REGION Network 14
   RUNG wire#powerrail
      #"2#柴油泵电动阀"(READY := "2#柴油泵电动蝶阀备妥", RUN := "2#柴油泵电动蝶阀运行", FAULT := "2#柴油泵电动蝶阀故障", OPEN_END := "2#柴油泵电动蝶阀开到位", CLOSE_END := "2#柴油泵电动蝶阀关到位", HMI_OPEN :=, HMI_CLOSE :=, MA :=, AUTO_OPEN :=, AUTO_CLOSE :=, QD_OPEN := "2#柴油泵电动阀开", QD_CLOSE := "2#柴油泵电动阀关")
   END_RUNG
   // the same network as SCL:
   #"2#柴油泵电动阀"(READY := "2#柴油泵电动蝶阀备妥",   // "阀门_MODEL"
               RUN := "2#柴油泵电动蝶阀运行",
               FAULT := "2#柴油泵电动蝶阀故障",
               OPEN_END := "2#柴油泵电动蝶阀开到位",
               CLOSE_END := "2#柴油泵电动蝶阀关到位",
               QD_OPEN := "2#柴油泵电动阀开",
               QD_CLOSE := "2#柴油泵电动阀关");
END_REGION

REGION Network 15
   RUNG wire#powerrail
      #"1#浊环热水泵电动阀"(READY := "1#浊环热水电动蝶阀备妥", RUN := "1#浊环热水电动蝶阀运行", FAULT := "1#浊环热水电动蝶阀故障", OPEN_END := "1#浊环热水电动蝶阀开到位", CLOSE_END := "1#浊环热水电动蝶阀关到位", HMI_OPEN :=, HMI_CLOSE :=, MA :=, AUTO_OPEN :=, AUTO_CLOSE :=, QD_OPEN := "1#浊环热水泵电动阀开", QD_CLOSE := "1#浊环热水泵电动阀关")
   END_RUNG
   // the same network as SCL:
   #"1#浊环热水泵电动阀"(READY := "1#浊环热水电动蝶阀备妥",   // "阀门_MODEL"
                 RUN := "1#浊环热水电动蝶阀运行",
                 FAULT := "1#浊环热水电动蝶阀故障",
                 OPEN_END := "1#浊环热水电动蝶阀开到位",
                 CLOSE_END := "1#浊环热水电动蝶阀关到位",
                 QD_OPEN := "1#浊环热水泵电动阀开",
                 QD_CLOSE := "1#浊环热水泵电动阀关");
END_REGION

REGION Network 16
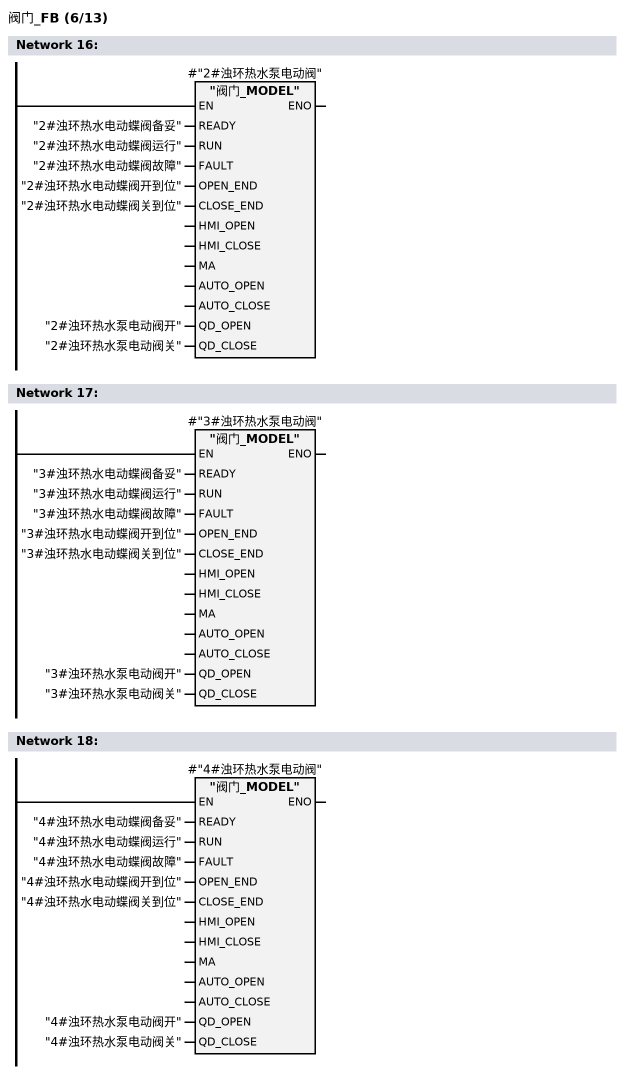
   RUNG wire#powerrail
      #"2#浊环热水泵电动阀"(READY := "2#浊环热水电动蝶阀备妥", RUN := "2#浊环热水电动蝶阀运行", FAULT := "2#浊环热水电动蝶阀故障", OPEN_END := "2#浊环热水电动蝶阀开到位", CLOSE_END := "2#浊环热水电动蝶阀关到位", HMI_OPEN :=, HMI_CLOSE :=, MA :=, AUTO_OPEN :=, AUTO_CLOSE :=, QD_OPEN := "2#浊环热水泵电动阀开", QD_CLOSE := "2#浊环热水泵电动阀关")
   END_RUNG
   // the same network as SCL:
   #"2#浊环热水泵电动阀"(READY := "2#浊环热水电动蝶阀备妥",   // "阀门_MODEL"
                 RUN := "2#浊环热水电动蝶阀运行",
                 FAULT := "2#浊环热水电动蝶阀故障",
                 OPEN_END := "2#浊环热水电动蝶阀开到位",
                 CLOSE_END := "2#浊环热水电动蝶阀关到位",
                 QD_OPEN := "2#浊环热水泵电动阀开",
                 QD_CLOSE := "2#浊环热水泵电动阀关");
END_REGION

REGION Network 17
   RUNG wire#powerrail
      #"3#浊环热水泵电动阀"(READY := "3#浊环热水电动蝶阀备妥", RUN := "3#浊环热水电动蝶阀运行", FAULT := "3#浊环热水电动蝶阀故障", OPEN_END := "3#浊环热水电动蝶阀开到位", CLOSE_END := "3#浊环热水电动蝶阀关到位", HMI_OPEN :=, HMI_CLOSE :=, MA :=, AUTO_OPEN :=, AUTO_CLOSE :=, QD_OPEN := "3#浊环热水泵电动阀开", QD_CLOSE := "3#浊环热水泵电动阀关")
   END_RUNG
   // the same network as SCL:
   #"3#浊环热水泵电动阀"(READY := "3#浊环热水电动蝶阀备妥",   // "阀门_MODEL"
                 RUN := "3#浊环热水电动蝶阀运行",
                 FAULT := "3#浊环热水电动蝶阀故障",
                 OPEN_END := "3#浊环热水电动蝶阀开到位",
                 CLOSE_END := "3#浊环热水电动蝶阀关到位",
                 QD_OPEN := "3#浊环热水泵电动阀开",
                 QD_CLOSE := "3#浊环热水泵电动阀关");
END_REGION

REGION Network 18
   RUNG wire#powerrail
      #"4#浊环热水泵电动阀"(READY := "4#浊环热水电动蝶阀备妥", RUN := "4#浊环热水电动蝶阀运行", FAULT := "4#浊环热水电动蝶阀故障", OPEN_END := "4#浊环热水电动蝶阀开到位", CLOSE_END := "4#浊环热水电动蝶阀关到位", HMI_OPEN :=, HMI_CLOSE :=, MA :=, AUTO_OPEN :=, AUTO_CLOSE :=, QD_OPEN := "4#浊环热水泵电动阀开", QD_CLOSE := "4#浊环热水泵电动阀关")
   END_RUNG
   // the same network as SCL:
   #"4#浊环热水泵电动阀"(READY := "4#浊环热水电动蝶阀备妥",   // "阀门_MODEL"
                 RUN := "4#浊环热水电动蝶阀运行",
                 FAULT := "4#浊环热水电动蝶阀故障",
                 OPEN_END := "4#浊环热水电动蝶阀开到位",
                 CLOSE_END := "4#浊环热水电动蝶阀关到位",
                 QD_OPEN := "4#浊环热水泵电动阀开",
                 QD_CLOSE := "4#浊环热水泵电动阀关");
END_REGION

REGION Network 19
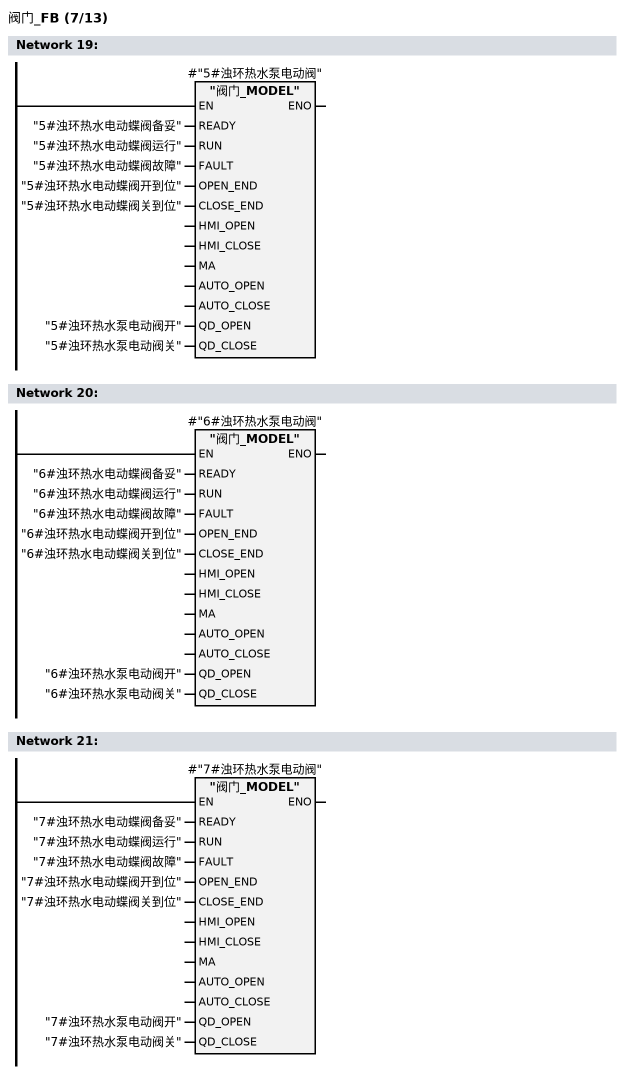
   RUNG wire#powerrail
      #"5#浊环热水泵电动阀"(READY := "5#浊环热水电动蝶阀备妥", RUN := "5#浊环热水电动蝶阀运行", FAULT := "5#浊环热水电动蝶阀故障", OPEN_END := "5#浊环热水电动蝶阀开到位", CLOSE_END := "5#浊环热水电动蝶阀关到位", HMI_OPEN :=, HMI_CLOSE :=, MA :=, AUTO_OPEN :=, AUTO_CLOSE :=, QD_OPEN := "5#浊环热水泵电动阀开", QD_CLOSE := "5#浊环热水泵电动阀关")
   END_RUNG
   // the same network as SCL:
   #"5#浊环热水泵电动阀"(READY := "5#浊环热水电动蝶阀备妥",   // "阀门_MODEL"
                 RUN := "5#浊环热水电动蝶阀运行",
                 FAULT := "5#浊环热水电动蝶阀故障",
                 OPEN_END := "5#浊环热水电动蝶阀开到位",
                 CLOSE_END := "5#浊环热水电动蝶阀关到位",
                 QD_OPEN := "5#浊环热水泵电动阀开",
                 QD_CLOSE := "5#浊环热水泵电动阀关");
END_REGION

REGION Network 20
   RUNG wire#powerrail
      #"6#浊环热水泵电动阀"(READY := "6#浊环热水电动蝶阀备妥", RUN := "6#浊环热水电动蝶阀运行", FAULT := "6#浊环热水电动蝶阀故障", OPEN_END := "6#浊环热水电动蝶阀开到位", CLOSE_END := "6#浊环热水电动蝶阀关到位", HMI_OPEN :=, HMI_CLOSE :=, MA :=, AUTO_OPEN :=, AUTO_CLOSE :=, QD_OPEN := "6#浊环热水泵电动阀开", QD_CLOSE := "6#浊环热水泵电动阀关")
   END_RUNG
   // the same network as SCL:
   #"6#浊环热水泵电动阀"(READY := "6#浊环热水电动蝶阀备妥",   // "阀门_MODEL"
                 RUN := "6#浊环热水电动蝶阀运行",
                 FAULT := "6#浊环热水电动蝶阀故障",
                 OPEN_END := "6#浊环热水电动蝶阀开到位",
                 CLOSE_END := "6#浊环热水电动蝶阀关到位",
                 QD_OPEN := "6#浊环热水泵电动阀开",
                 QD_CLOSE := "6#浊环热水泵电动阀关");
END_REGION

REGION Network 21
   RUNG wire#powerrail
      #"7#浊环热水泵电动阀"(READY := "7#浊环热水电动蝶阀备妥", RUN := "7#浊环热水电动蝶阀运行", FAULT := "7#浊环热水电动蝶阀故障", OPEN_END := "7#浊环热水电动蝶阀开到位", CLOSE_END := "7#浊环热水电动蝶阀关到位", HMI_OPEN :=, HMI_CLOSE :=, MA :=, AUTO_OPEN :=, AUTO_CLOSE :=, QD_OPEN := "7#浊环热水泵电动阀开", QD_CLOSE := "7#浊环热水泵电动阀关")
   END_RUNG
   // the same network as SCL:
   #"7#浊环热水泵电动阀"(READY := "7#浊环热水电动蝶阀备妥",   // "阀门_MODEL"
                 RUN := "7#浊环热水电动蝶阀运行",
                 FAULT := "7#浊环热水电动蝶阀故障",
                 OPEN_END := "7#浊环热水电动蝶阀开到位",
                 CLOSE_END := "7#浊环热水电动蝶阀关到位",
                 QD_OPEN := "7#浊环热水泵电动阀开",
                 QD_CLOSE := "7#浊环热水泵电动阀关");
END_REGION

REGION Network 22
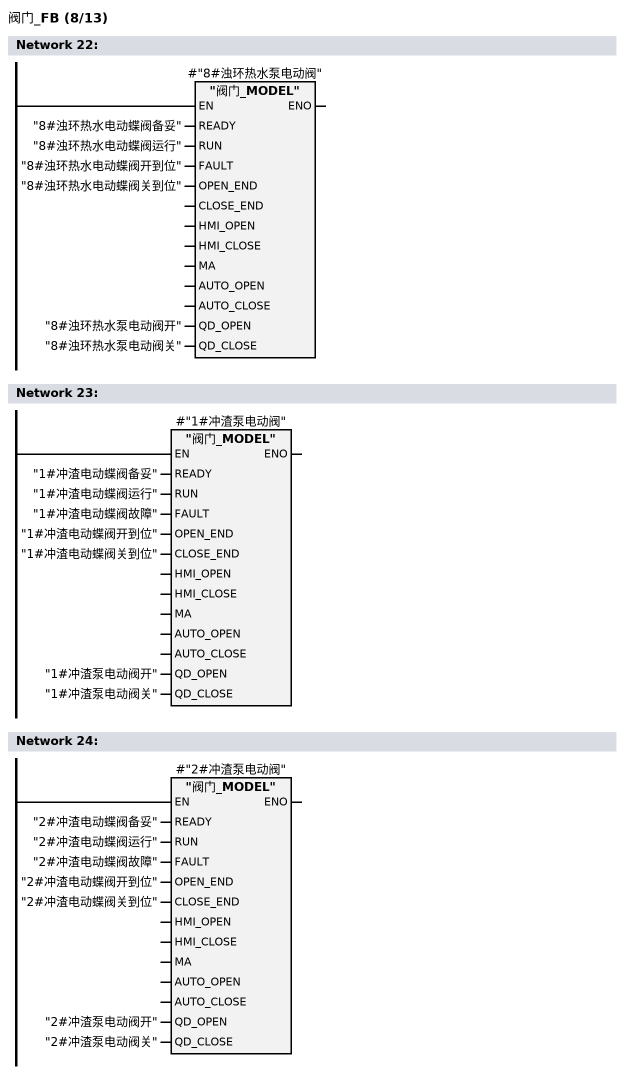
   RUNG wire#powerrail
      #"8#浊环热水泵电动阀"(READY := "8#浊环热水电动蝶阀备妥", RUN := "8#浊环热水电动蝶阀运行", FAULT := "8#浊环热水电动蝶阀开到位", OPEN_END := "8#浊环热水电动蝶阀关到位", CLOSE_END :=, HMI_OPEN :=, HMI_CLOSE :=, MA :=, AUTO_OPEN :=, AUTO_CLOSE :=, QD_OPEN := "8#浊环热水泵电动阀开", QD_CLOSE := "8#浊环热水泵电动阀关")
   END_RUNG
   // the same network as SCL:
   #"8#浊环热水泵电动阀"(READY := "8#浊环热水电动蝶阀备妥",   // "阀门_MODEL"
                 RUN := "8#浊环热水电动蝶阀运行",
                 FAULT := "8#浊环热水电动蝶阀开到位",
                 OPEN_END := "8#浊环热水电动蝶阀关到位",
                 QD_OPEN := "8#浊环热水泵电动阀开",
                 QD_CLOSE := "8#浊环热水泵电动阀关");
END_REGION

REGION Network 23
   RUNG wire#powerrail
      #"1#冲渣泵电动阀"(READY := "1#冲渣电动蝶阀备妥", RUN := "1#冲渣电动蝶阀运行", FAULT := "1#冲渣电动蝶阀故障", OPEN_END := "1#冲渣电动蝶阀开到位", CLOSE_END := "1#冲渣电动蝶阀关到位", HMI_OPEN :=, HMI_CLOSE :=, MA :=, AUTO_OPEN :=, AUTO_CLOSE :=, QD_OPEN := "1#冲渣泵电动阀开", QD_CLOSE := "1#冲渣泵电动阀关")
   END_RUNG
   // the same network as SCL:
   #"1#冲渣泵电动阀"(READY := "1#冲渣电动蝶阀备妥",   // "阀门_MODEL"
               RUN := "1#冲渣电动蝶阀运行",
               FAULT := "1#冲渣电动蝶阀故障",
               OPEN_END := "1#冲渣电动蝶阀开到位",
               CLOSE_END := "1#冲渣电动蝶阀关到位",
               QD_OPEN := "1#冲渣泵电动阀开",
               QD_CLOSE := "1#冲渣泵电动阀关");
END_REGION

REGION Network 24
   RUNG wire#powerrail
      #"2#冲渣泵电动阀"(READY := "2#冲渣电动蝶阀备妥", RUN := "2#冲渣电动蝶阀运行", FAULT := "2#冲渣电动蝶阀故障", OPEN_END := "2#冲渣电动蝶阀开到位", CLOSE_END := "2#冲渣电动蝶阀关到位", HMI_OPEN :=, HMI_CLOSE :=, MA :=, AUTO_OPEN :=, AUTO_CLOSE :=, QD_OPEN := "2#冲渣泵电动阀开", QD_CLOSE := "2#冲渣泵电动阀关")
   END_RUNG
   // the same network as SCL:
   #"2#冲渣泵电动阀"(READY := "2#冲渣电动蝶阀备妥",   // "阀门_MODEL"
               RUN := "2#冲渣电动蝶阀运行",
               FAULT := "2#冲渣电动蝶阀故障",
               OPEN_END := "2#冲渣电动蝶阀开到位",
               CLOSE_END := "2#冲渣电动蝶阀关到位",
               QD_OPEN := "2#冲渣泵电动阀开",
               QD_CLOSE := "2#冲渣泵电动阀关");
END_REGION

REGION Network 25
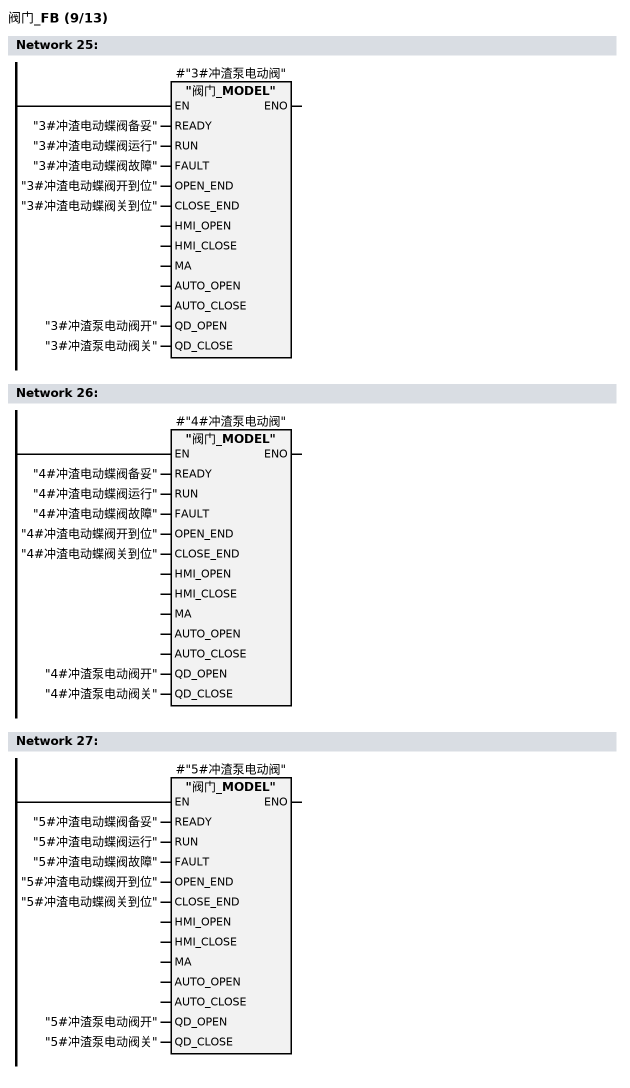
   RUNG wire#powerrail
      #"3#冲渣泵电动阀"(READY := "3#冲渣电动蝶阀备妥", RUN := "3#冲渣电动蝶阀运行", FAULT := "3#冲渣电动蝶阀故障", OPEN_END := "3#冲渣电动蝶阀开到位", CLOSE_END := "3#冲渣电动蝶阀关到位", HMI_OPEN :=, HMI_CLOSE :=, MA :=, AUTO_OPEN :=, AUTO_CLOSE :=, QD_OPEN := "3#冲渣泵电动阀开", QD_CLOSE := "3#冲渣泵电动阀关")
   END_RUNG
   // the same network as SCL:
   #"3#冲渣泵电动阀"(READY := "3#冲渣电动蝶阀备妥",   // "阀门_MODEL"
               RUN := "3#冲渣电动蝶阀运行",
               FAULT := "3#冲渣电动蝶阀故障",
               OPEN_END := "3#冲渣电动蝶阀开到位",
               CLOSE_END := "3#冲渣电动蝶阀关到位",
               QD_OPEN := "3#冲渣泵电动阀开",
               QD_CLOSE := "3#冲渣泵电动阀关");
END_REGION

REGION Network 26
   RUNG wire#powerrail
      #"4#冲渣泵电动阀"(READY := "4#冲渣电动蝶阀备妥", RUN := "4#冲渣电动蝶阀运行", FAULT := "4#冲渣电动蝶阀故障", OPEN_END := "4#冲渣电动蝶阀开到位", CLOSE_END := "4#冲渣电动蝶阀关到位", HMI_OPEN :=, HMI_CLOSE :=, MA :=, AUTO_OPEN :=, AUTO_CLOSE :=, QD_OPEN := "4#冲渣泵电动阀开", QD_CLOSE := "4#冲渣泵电动阀关")
   END_RUNG
   // the same network as SCL:
   #"4#冲渣泵电动阀"(READY := "4#冲渣电动蝶阀备妥",   // "阀门_MODEL"
               RUN := "4#冲渣电动蝶阀运行",
               FAULT := "4#冲渣电动蝶阀故障",
               OPEN_END := "4#冲渣电动蝶阀开到位",
               CLOSE_END := "4#冲渣电动蝶阀关到位",
               QD_OPEN := "4#冲渣泵电动阀开",
               QD_CLOSE := "4#冲渣泵电动阀关");
END_REGION

REGION Network 27
   RUNG wire#powerrail
      #"5#冲渣泵电动阀"(READY := "5#冲渣电动蝶阀备妥", RUN := "5#冲渣电动蝶阀运行", FAULT := "5#冲渣电动蝶阀故障", OPEN_END := "5#冲渣电动蝶阀开到位", CLOSE_END := "5#冲渣电动蝶阀关到位", HMI_OPEN :=, HMI_CLOSE :=, MA :=, AUTO_OPEN :=, AUTO_CLOSE :=, QD_OPEN := "5#冲渣泵电动阀开", QD_CLOSE := "5#冲渣泵电动阀关")
   END_RUNG
   // the same network as SCL:
   #"5#冲渣泵电动阀"(READY := "5#冲渣电动蝶阀备妥",   // "阀门_MODEL"
               RUN := "5#冲渣电动蝶阀运行",
               FAULT := "5#冲渣电动蝶阀故障",
               OPEN_END := "5#冲渣电动蝶阀开到位",
               CLOSE_END := "5#冲渣电动蝶阀关到位",
               QD_OPEN := "5#冲渣泵电动阀开",
               QD_CLOSE := "5#冲渣泵电动阀关");
END_REGION

REGION Network 28
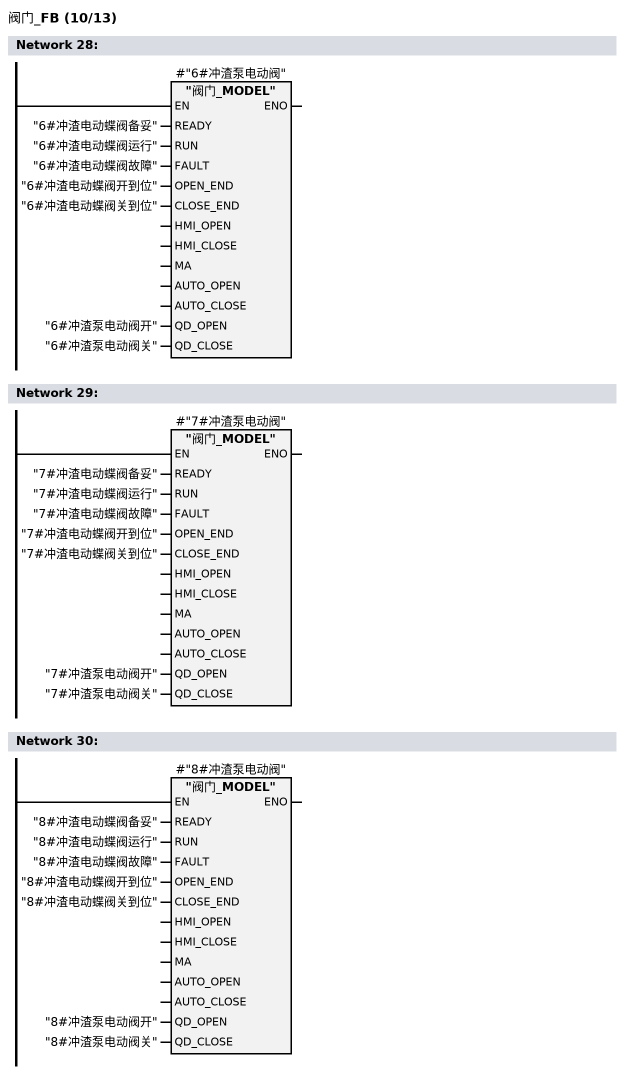
   RUNG wire#powerrail
      #"6#冲渣泵电动阀"(READY := "6#冲渣电动蝶阀备妥", RUN := "6#冲渣电动蝶阀运行", FAULT := "6#冲渣电动蝶阀故障", OPEN_END := "6#冲渣电动蝶阀开到位", CLOSE_END := "6#冲渣电动蝶阀关到位", HMI_OPEN :=, HMI_CLOSE :=, MA :=, AUTO_OPEN :=, AUTO_CLOSE :=, QD_OPEN := "6#冲渣泵电动阀开", QD_CLOSE := "6#冲渣泵电动阀关")
   END_RUNG
   // the same network as SCL:
   #"6#冲渣泵电动阀"(READY := "6#冲渣电动蝶阀备妥",   // "阀门_MODEL"
               RUN := "6#冲渣电动蝶阀运行",
               FAULT := "6#冲渣电动蝶阀故障",
               OPEN_END := "6#冲渣电动蝶阀开到位",
               CLOSE_END := "6#冲渣电动蝶阀关到位",
               QD_OPEN := "6#冲渣泵电动阀开",
               QD_CLOSE := "6#冲渣泵电动阀关");
END_REGION

REGION Network 29
   RUNG wire#powerrail
      #"7#冲渣泵电动阀"(READY := "7#冲渣电动蝶阀备妥", RUN := "7#冲渣电动蝶阀运行", FAULT := "7#冲渣电动蝶阀故障", OPEN_END := "7#冲渣电动蝶阀开到位", CLOSE_END := "7#冲渣电动蝶阀关到位", HMI_OPEN :=, HMI_CLOSE :=, MA :=, AUTO_OPEN :=, AUTO_CLOSE :=, QD_OPEN := "7#冲渣泵电动阀开", QD_CLOSE := "7#冲渣泵电动阀关")
   END_RUNG
   // the same network as SCL:
   #"7#冲渣泵电动阀"(READY := "7#冲渣电动蝶阀备妥",   // "阀门_MODEL"
               RUN := "7#冲渣电动蝶阀运行",
               FAULT := "7#冲渣电动蝶阀故障",
               OPEN_END := "7#冲渣电动蝶阀开到位",
               CLOSE_END := "7#冲渣电动蝶阀关到位",
               QD_OPEN := "7#冲渣泵电动阀开",
               QD_CLOSE := "7#冲渣泵电动阀关");
END_REGION

REGION Network 30
   RUNG wire#powerrail
      #"8#冲渣泵电动阀"(READY := "8#冲渣电动蝶阀备妥", RUN := "8#冲渣电动蝶阀运行", FAULT := "8#冲渣电动蝶阀故障", OPEN_END := "8#冲渣电动蝶阀开到位", CLOSE_END := "8#冲渣电动蝶阀关到位", HMI_OPEN :=, HMI_CLOSE :=, MA :=, AUTO_OPEN :=, AUTO_CLOSE :=, QD_OPEN := "8#冲渣泵电动阀开", QD_CLOSE := "8#冲渣泵电动阀关")
   END_RUNG
   // the same network as SCL:
   #"8#冲渣泵电动阀"(READY := "8#冲渣电动蝶阀备妥",   // "阀门_MODEL"
               RUN := "8#冲渣电动蝶阀运行",
               FAULT := "8#冲渣电动蝶阀故障",
               OPEN_END := "8#冲渣电动蝶阀开到位",
               CLOSE_END := "8#冲渣电动蝶阀关到位",
               QD_OPEN := "8#冲渣泵电动阀开",
               QD_CLOSE := "8#冲渣泵电动阀关");
END_REGION

REGION Network 31
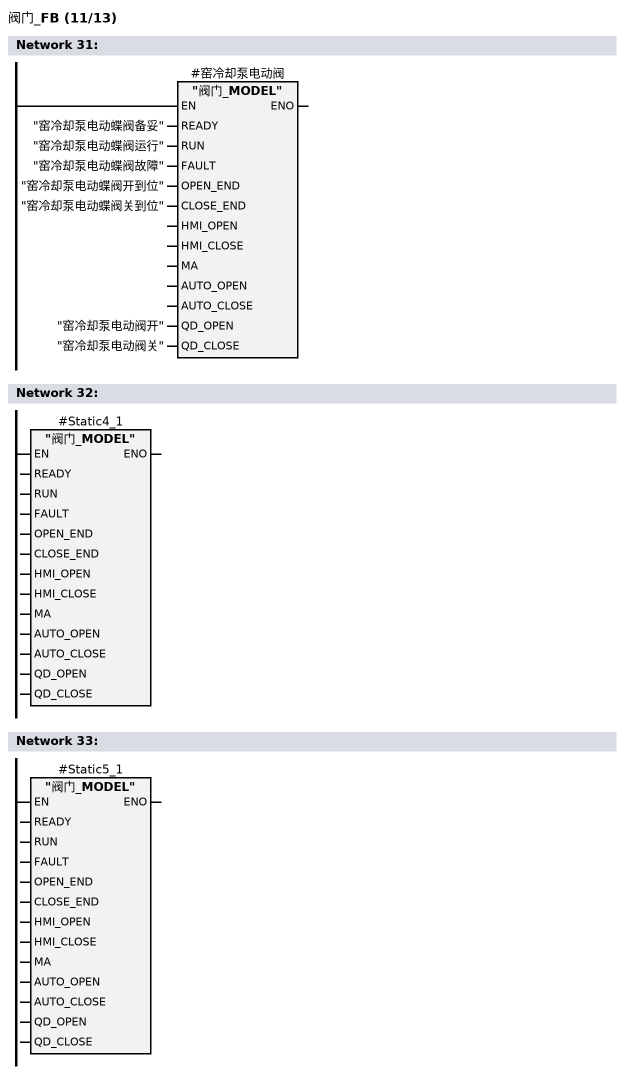
   RUNG wire#powerrail
      #窑冷却泵电动阀(READY := "窑冷却泵电动蝶阀备妥", RUN := "窑冷却泵电动蝶阀运行", FAULT := "窑冷却泵电动蝶阀故障", OPEN_END := "窑冷却泵电动蝶阀开到位", CLOSE_END := "窑冷却泵电动蝶阀关到位", HMI_OPEN :=, HMI_CLOSE :=, MA :=, AUTO_OPEN :=, AUTO_CLOSE :=, QD_OPEN := "窑冷却泵电动阀开", QD_CLOSE := "窑冷却泵电动阀关")
   END_RUNG
   // the same network as SCL:
   #窑冷却泵电动阀(READY := "窑冷却泵电动蝶阀备妥",   // "阀门_MODEL"
            RUN := "窑冷却泵电动蝶阀运行",
            FAULT := "窑冷却泵电动蝶阀故障",
            OPEN_END := "窑冷却泵电动蝶阀开到位",
            CLOSE_END := "窑冷却泵电动蝶阀关到位",
            QD_OPEN := "窑冷却泵电动阀开",
            QD_CLOSE := "窑冷却泵电动阀关");
END_REGION

REGION Network 32
   RUNG wire#powerrail
      #Static4_1(READY :=, RUN :=, FAULT :=, OPEN_END :=, CLOSE_END :=, HMI_OPEN :=, HMI_CLOSE :=, MA :=, AUTO_OPEN :=, AUTO_CLOSE :=, QD_OPEN :=, QD_CLOSE :=)
   END_RUNG
   // the same network as SCL:
   #Static4_1();   // "阀门_MODEL"
END_REGION

REGION Network 33
   RUNG wire#powerrail
      #Static5_1(READY :=, RUN :=, FAULT :=, OPEN_END :=, CLOSE_END :=, HMI_OPEN :=, HMI_CLOSE :=, MA :=, AUTO_OPEN :=, AUTO_CLOSE :=, QD_OPEN :=, QD_CLOSE :=)
   END_RUNG
   // the same network as SCL:
   #Static5_1();   // "阀门_MODEL"
END_REGION

REGION Network 34
